REGION Network 7: Send Current Mode
   // Relay current mode to master & slave
   RUNG wire#powerrail
      Move(in := "70_Mode_Data".CRNT_MODE, out1 => "56_SLAVE_CMNDS".CRNT_MODE)
      Move(in := "70_Mode_Data".CRNT_MODE, out1 => "55_STATUS_DATA".CRNT_MODE)
      Move(in := "70_Mode_Data".CRNT_MODE, out1 => "82_To_HMI".CRNT_MODE_IGG)
   END_RUNG
   // the same network as SCL:
   "56_SLAVE_CMNDS".CRNT_MODE := "70_Mode_Data".CRNT_MODE;
   "55_STATUS_DATA".CRNT_MODE := "70_Mode_Data".CRNT_MODE;
   "82_To_HMI".CRNT_MODE_IGG := "70_Mode_Data".CRNT_MODE;
END_REGION

REGION Network 8: Leaving Manual
   // For determination of transition to automatic
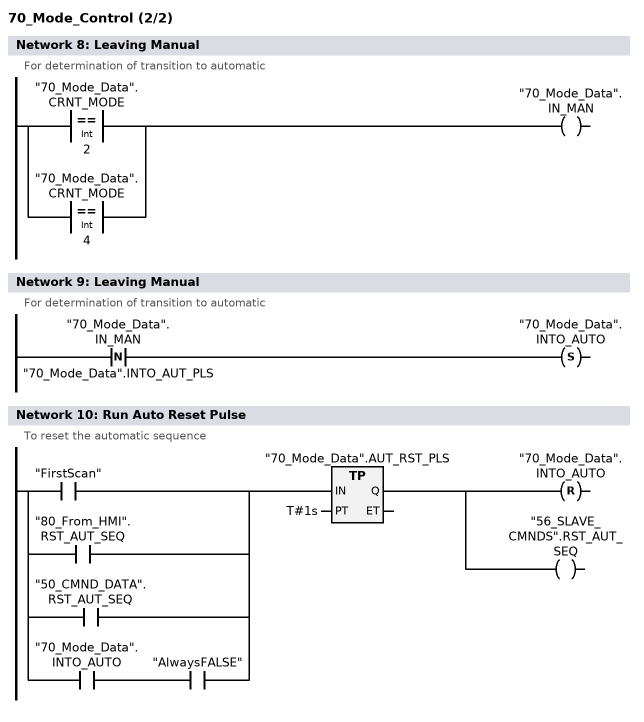
   RUNG wire#powerrail
      { S7_Templates := "SrcType := Int" } EQ_Contact(in1 := "70_Mode_Data".CRNT_MODE, in2 := 2)
      wire#w1
      Coil( "70_Mode_Data".IN_MAN )
   END_RUNG
   RUNG wire#powerrail
      { S7_Templates := "SrcType := Int" } EQ_Contact(in1 := "70_Mode_Data".CRNT_MODE, in2 := 4)
   END_RUNG wire#w1
   // the same network as SCL:
   "70_Mode_Data".IN_MAN := ("70_Mode_Data".CRNT_MODE = 2) OR ("70_Mode_Data".CRNT_MODE = 4);
END_REGION

REGION Network 9: Leaving Manual
   // For determination of transition to automatic
   RUNG wire#powerrail
      N_Contact(operand := "70_Mode_Data".IN_MAN, bit := "70_Mode_Data".INTO_AUT_PLS)
      S_Coil( "70_Mode_Data".INTO_AUTO )
   END_RUNG
   // the same network as SCL:
   #_w1 := NOT "70_Mode_Data".IN_MAN AND "70_Mode_Data".INTO_AUT_PLS;   // falling edge of "70_Mode_Data".IN_MAN
   "70_Mode_Data".INTO_AUT_PLS := "70_Mode_Data".IN_MAN;
   IF #_w1 THEN "70_Mode_Data".INTO_AUTO := TRUE; END_IF;
END_REGION

REGION Network 10: Run Auto Reset Pulse
   // To reset the automatic sequence
   "70_Mode_Data".AUT_RST_PLS.TP(IN := "FirstScan" OR "80_From_HMI".RST_AUT_SEQ OR "50_CMND_DATA".RST_AUT_SEQ OR ("70_Mode_Data".INTO_AUTO AND "AlwaysFALSE"),
                           PT := T#1s);
   IF "70_Mode_Data".AUT_RST_PLS.Q THEN "70_Mode_Data".INTO_AUTO := FALSE; END_IF;
   "56_SLAVE_CMNDS".RST_AUT_SEQ := "70_Mode_Data".AUT_RST_PLS.Q;
END_REGION
END_FUNCTION

// folder: 90 - 99 Manual Functions

FUNCTION_BLOCK "FuelPump"   // FB505, LAD
{ S7_Optimized_Access := 'TRUE' }
VERSION : 0.1
   VAR_INPUT
      Start_Command : Bool;
      Triped : Bool;
      Run : Bool;
      "E-Stop" : Bool;
      Interlock : Bool;
   END_VAR
   VAR_OUTPUT
      Start_Pump : Bool;
   END_VAR
   VAR
      Aux : Struct
         Aux1 : Bool;
         Aux2 : Bool;
      END_STRUCT;
   END_VAR
   VAR_TEMP   // added for the SCL form of the ladder/FBD networks
      _w1 : Bool;
      _w2 : Bool;
      _w3 : Bool;
   END_VAR
BEGIN

REGION Network 1
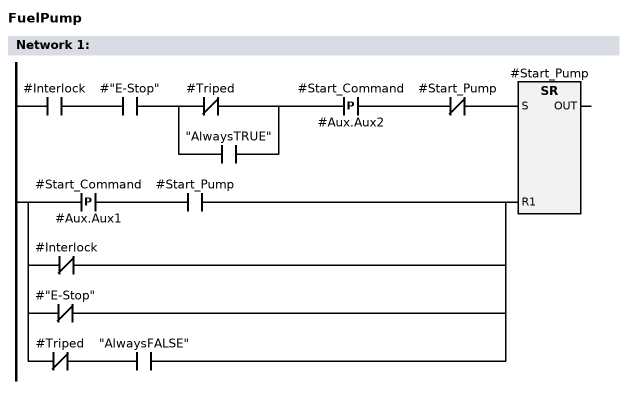
   RUNG wire#powerrail
      Contact( #Interlock )
      Contact( #"E-Stop" )
      wire#w1
      I_Contact( #Triped )
      wire#w2
      P_Contact(operand := #Start_Command, bit := #Aux.Aux2)
      I_Contact( #Start_Pump )
      S_SR(operand := #Start_Pump, r1 := wire#w3)
   END_RUNG
   RUNG wire#w1
      Contact( "AlwaysTRUE" )
   END_RUNG wire#w2
   RUNG wire#powerrail
      P_Contact(operand := #Start_Command, bit := #Aux.Aux1)
      Contact( #Start_Pump )
   END_RUNG wire#w3
   RUNG wire#powerrail
      I_Contact( #Interlock )
   END_RUNG wire#w3
   RUNG wire#powerrail
      I_Contact( #"E-Stop" )
   END_RUNG wire#w3
   RUNG wire#powerrail
      I_Contact( #Triped )
      Contact( "AlwaysFALSE" )
   END_RUNG wire#w3
   // the same network as SCL:
   #_w1 := #Interlock AND #"E-Stop" AND (NOT #Triped OR "AlwaysTRUE") AND #Start_Command AND NOT #Aux.Aux2;   // rising edge of #Start_Command
   #Aux.Aux2 := #Start_Command;
   #_w2 := #Start_Command AND NOT #Aux.Aux1;   // rising edge of #Start_Command
   #Aux.Aux1 := #Start_Command;
   #_w3 := (#_w2 AND #Start_Pump) OR NOT #Interlock OR NOT #"E-Stop" OR (NOT #Triped AND "AlwaysFALSE");
   IF #_w1 AND NOT #Start_Pump THEN
       #Start_Pump := TRUE;   // SR flip-flop
   END_IF;
   IF #_w3 THEN #Start_Pump := FALSE; END_IF;
END_REGION
END_FUNCTION_BLOCK

FUNCTION "90_Manual_Control" : Void   // FC90, LAD
TITLE = Manual Control
{ S7_Optimized_Access := 'TRUE' }
AUTHOR : JHT
VERSION : 0.1
// Code for manual operation of equipment
   VAR_TEMP
      Aux : Struct
         Aux1 : Bool;
      END_STRUCT;
   END_VAR
   VAR_TEMP   // added for the SCL form of the ladder/FBD networks
      _w1 : Bool;
      _w2 : Bool;
      _w3 : Bool;
      _w4 : Bool;
      _w5 : Bool;
      _w6 : Bool;
   END_VAR
BEGIN

REGION Network 1: Zero Auto Step Numbers
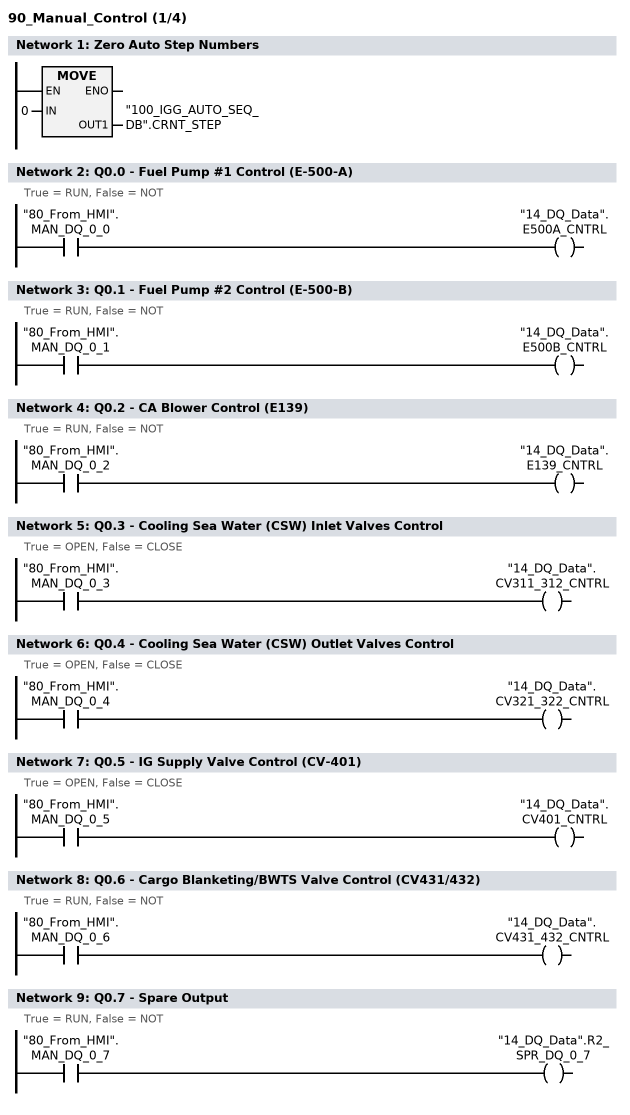
   RUNG wire#powerrail
      Move(in := 0, out1 => "100_IGG_AUTO_SEQ_DB".CRNT_STEP)
   END_RUNG
   // the same network as SCL:
   "100_IGG_AUTO_SEQ_DB".CRNT_STEP := 0;
END_REGION

REGION Network 2: Q0.0 - Fuel Pump #1 Control (E-500-A)
   // True = RUN, False = NOT
   RUNG wire#powerrail
      Contact( "80_From_HMI".MAN_DQ_0_0 )
      Coil( "14_DQ_Data".E500A_CNTRL )
   END_RUNG
   // the same network as SCL:
   "14_DQ_Data".E500A_CNTRL := "80_From_HMI".MAN_DQ_0_0;
END_REGION

REGION Network 3: Q0.1 - Fuel Pump #2 Control (E-500-B)
   // True = RUN, False = NOT
   RUNG wire#powerrail
      Contact( "80_From_HMI".MAN_DQ_0_1 )
      Coil( "14_DQ_Data".E500B_CNTRL )
   END_RUNG
   // the same network as SCL:
   "14_DQ_Data".E500B_CNTRL := "80_From_HMI".MAN_DQ_0_1;
END_REGION

REGION Network 4: Q0.2 - CA Blower Control (E139)
   // True = RUN, False = NOT
   RUNG wire#powerrail
      Contact( "80_From_HMI".MAN_DQ_0_2 )
      Coil( "14_DQ_Data".E139_CNTRL )
   END_RUNG
   // the same network as SCL:
   "14_DQ_Data".E139_CNTRL := "80_From_HMI".MAN_DQ_0_2;
END_REGION

REGION Network 5: Q0.3 - Cooling Sea Water (CSW) Inlet Valves Control
   // True = OPEN, False = CLOSE
   RUNG wire#powerrail
      Contact( "80_From_HMI".MAN_DQ_0_3 )
      Coil( "14_DQ_Data".CV311_312_CNTRL )
   END_RUNG
   // the same network as SCL:
   "14_DQ_Data".CV311_312_CNTRL := "80_From_HMI".MAN_DQ_0_3;
END_REGION

REGION Network 6: Q0.4 - Cooling Sea Water (CSW) Outlet Valves Control
   // True = OPEN, False = CLOSE
   RUNG wire#powerrail
      Contact( "80_From_HMI".MAN_DQ_0_4 )
      Coil( "14_DQ_Data".CV321_322_CNTRL )
   END_RUNG
   // the same network as SCL:
   "14_DQ_Data".CV321_322_CNTRL := "80_From_HMI".MAN_DQ_0_4;
END_REGION

REGION Network 7: Q0.5 - IG Supply Valve Control (CV-401)
   // True = OPEN, False = CLOSE
   RUNG wire#powerrail
      Contact( "80_From_HMI".MAN_DQ_0_5 )
      Coil( "14_DQ_Data".CV401_CNTRL )
   END_RUNG
   // the same network as SCL:
   "14_DQ_Data".CV401_CNTRL := "80_From_HMI".MAN_DQ_0_5;
END_REGION

REGION Network 8: Q0.6 - Cargo Blanketing/BWTS Valve Control (CV431/432)
   // True = RUN, False = NOT
   RUNG wire#powerrail
      Contact( "80_From_HMI".MAN_DQ_0_6 )
      Coil( "14_DQ_Data".CV431_432_CNTRL )
   END_RUNG
   // the same network as SCL:
   "14_DQ_Data".CV431_432_CNTRL := "80_From_HMI".MAN_DQ_0_6;
END_REGION

REGION Network 9: Q0.7 - Spare Output
   // True = RUN, False = NOT
   RUNG wire#powerrail
      Contact( "80_From_HMI".MAN_DQ_0_7 )
      Coil( "14_DQ_Data".R2_SPR_DQ_0_7 )
   END_RUNG
   // the same network as SCL:
   "14_DQ_Data".R2_SPR_DQ_0_7 := "80_From_HMI".MAN_DQ_0_7;
END_REGION

REGION Network 10: Q1.0 - Spare Output
   // True = RUN, False = NOT
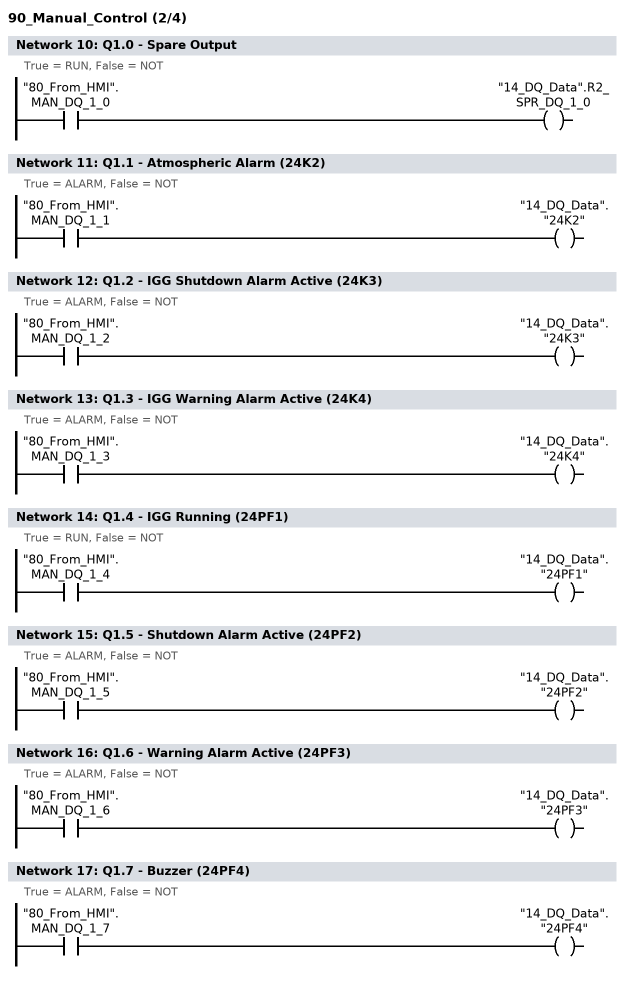
   RUNG wire#powerrail
      Contact( "80_From_HMI".MAN_DQ_1_0 )
      Coil( "14_DQ_Data".R2_SPR_DQ_1_0 )
   END_RUNG
   // the same network as SCL:
   "14_DQ_Data".R2_SPR_DQ_1_0 := "80_From_HMI".MAN_DQ_1_0;
END_REGION

REGION Network 11: Q1.1 - Atmospheric Alarm (24K2)
   // True = ALARM, False = NOT
   RUNG wire#powerrail
      Contact( "80_From_HMI".MAN_DQ_1_1 )
      Coil( "14_DQ_Data"."24K2" )
   END_RUNG
   // the same network as SCL:
   "14_DQ_Data"."24K2" := "80_From_HMI".MAN_DQ_1_1;
END_REGION

REGION Network 12: Q1.2 - IGG Shutdown Alarm Active (24K3)
   // True = ALARM, False = NOT
   RUNG wire#powerrail
      Contact( "80_From_HMI".MAN_DQ_1_2 )
      Coil( "14_DQ_Data"."24K3" )
   END_RUNG
   // the same network as SCL:
   "14_DQ_Data"."24K3" := "80_From_HMI".MAN_DQ_1_2;
END_REGION

REGION Network 13: Q1.3 - IGG Warning Alarm Active (24K4)
   // True = ALARM, False = NOT
   RUNG wire#powerrail
      Contact( "80_From_HMI".MAN_DQ_1_3 )
      Coil( "14_DQ_Data"."24K4" )
   END_RUNG
   // the same network as SCL:
   "14_DQ_Data"."24K4" := "80_From_HMI".MAN_DQ_1_3;
END_REGION

REGION Network 14: Q1.4 - IGG Running (24PF1)
   // True = RUN, False = NOT
   RUNG wire#powerrail
      Contact( "80_From_HMI".MAN_DQ_1_4 )
      Coil( "14_DQ_Data"."24PF1" )
   END_RUNG
   // the same network as SCL:
   "14_DQ_Data"."24PF1" := "80_From_HMI".MAN_DQ_1_4;
END_REGION

REGION Network 15: Q1.5 - Shutdown Alarm Active (24PF2)
   // True = ALARM, False = NOT
   RUNG wire#powerrail
      Contact( "80_From_HMI".MAN_DQ_1_5 )
      Coil( "14_DQ_Data"."24PF2" )
   END_RUNG
   // the same network as SCL:
   "14_DQ_Data"."24PF2" := "80_From_HMI".MAN_DQ_1_5;
END_REGION

REGION Network 16: Q1.6 - Warning Alarm Active (24PF3)
   // True = ALARM, False = NOT
   RUNG wire#powerrail
      Contact( "80_From_HMI".MAN_DQ_1_6 )
      Coil( "14_DQ_Data"."24PF3" )
   END_RUNG
   // the same network as SCL:
   "14_DQ_Data"."24PF3" := "80_From_HMI".MAN_DQ_1_6;
END_REGION

REGION Network 17: Q1.7 - Buzzer (24PF4)
   // True = ALARM, False = NOT
   RUNG wire#powerrail
      Contact( "80_From_HMI".MAN_DQ_1_7 )
      Coil( "14_DQ_Data"."24PF4" )
   END_RUNG
   // the same network as SCL:
   "14_DQ_Data"."24PF4" := "80_From_HMI".MAN_DQ_1_7;
END_REGION

REGION Network 18: QW98 - Vent Valve Position Control (CV-403)
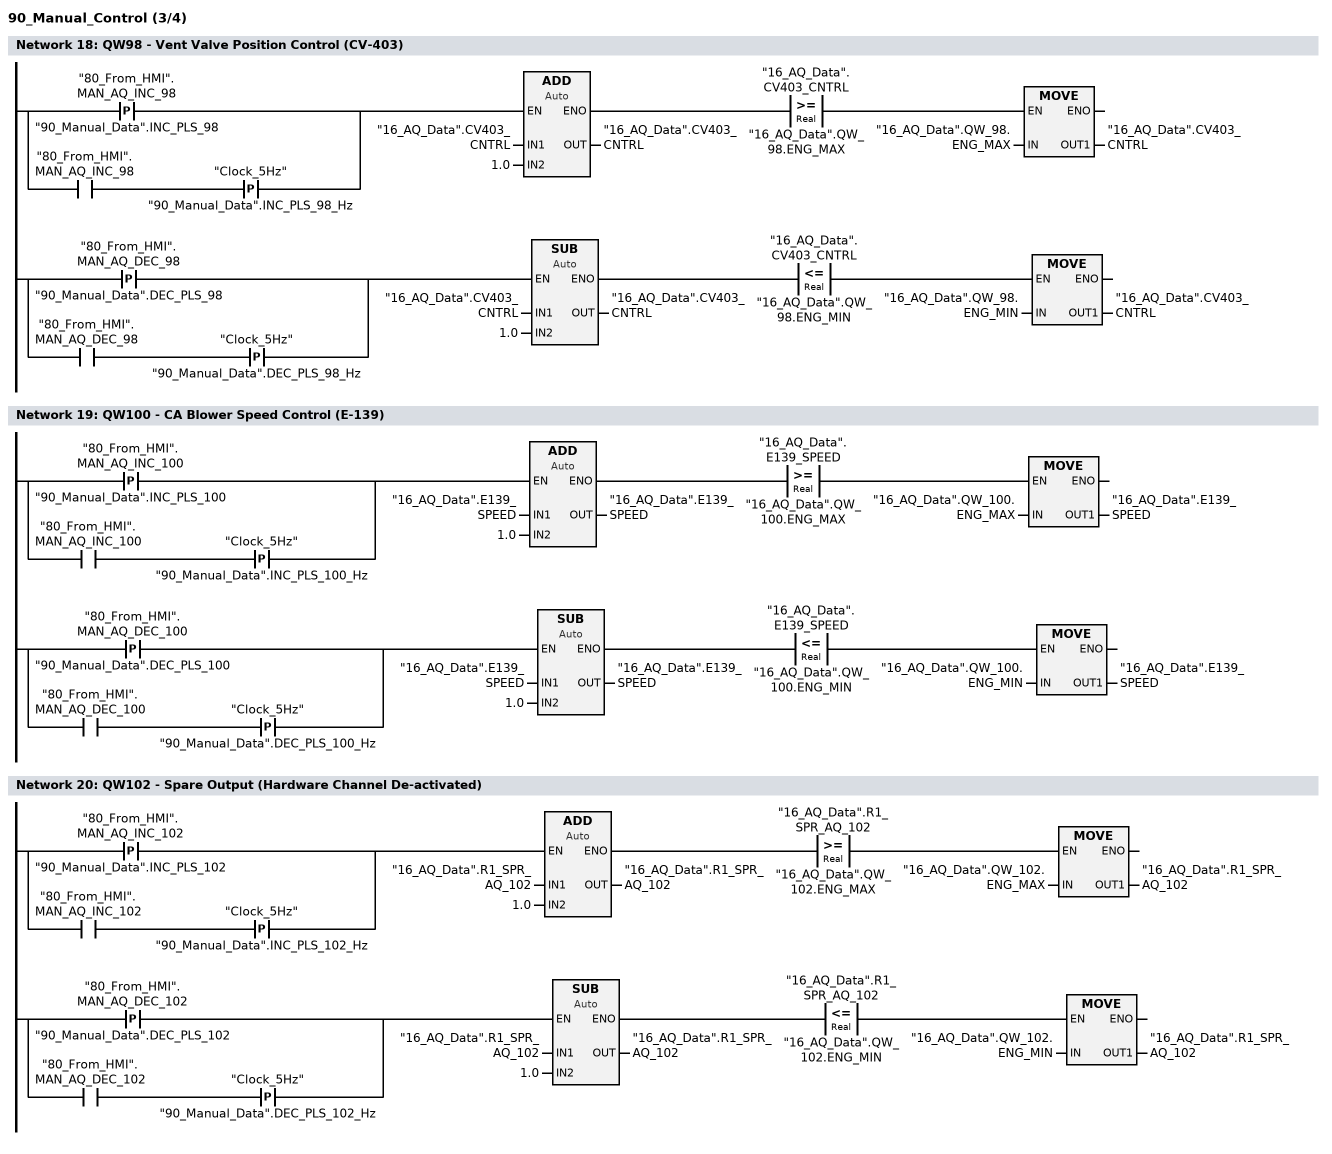
   RUNG wire#powerrail
      P_Contact(operand := "80_From_HMI".MAN_AQ_INC_98, bit := "90_Manual_Data".INC_PLS_98)
      wire#w1
      Add(in1 := "16_AQ_Data".CV403_CNTRL, in2 := 1.0, out => "16_AQ_Data".CV403_CNTRL)
      { S7_Templates := "SrcType := Real" } GE_Contact(in1 := "16_AQ_Data".CV403_CNTRL, in2 := "16_AQ_Data".QW_98.ENG_MAX)
      { S7_GenerateENO := "TRUE" } Move(in := "16_AQ_Data".QW_98.ENG_MAX, out1 => "16_AQ_Data".CV403_CNTRL)
   END_RUNG
   RUNG wire#powerrail
      Contact( "80_From_HMI".MAN_AQ_INC_98 )
      P_Contact(operand := "Clock_5Hz", bit := "90_Manual_Data".INC_PLS_98_Hz)
   END_RUNG wire#w1
   RUNG wire#powerrail
      P_Contact(operand := "80_From_HMI".MAN_AQ_DEC_98, bit := "90_Manual_Data".DEC_PLS_98)
      wire#w2
      Sub(in1 := "16_AQ_Data".CV403_CNTRL, in2 := 1.0, out => "16_AQ_Data".CV403_CNTRL)
      { S7_Templates := "SrcType := Real" } LE_Contact(in1 := "16_AQ_Data".CV403_CNTRL, in2 := "16_AQ_Data".QW_98.ENG_MIN)
      { S7_GenerateENO := "TRUE" } Move(in := "16_AQ_Data".QW_98.ENG_MIN, out1 => "16_AQ_Data".CV403_CNTRL)
   END_RUNG
   RUNG wire#powerrail
      Contact( "80_From_HMI".MAN_AQ_DEC_98 )
      P_Contact(operand := "Clock_5Hz", bit := "90_Manual_Data".DEC_PLS_98_Hz)
   END_RUNG wire#w2
   // the same network as SCL:
   #_w1 := "80_From_HMI".MAN_AQ_INC_98 AND NOT "90_Manual_Data".INC_PLS_98;   // rising edge of "80_From_HMI".MAN_AQ_INC_98
   "90_Manual_Data".INC_PLS_98 := "80_From_HMI".MAN_AQ_INC_98;
   #_w2 := "80_From_HMI".MAN_AQ_INC_98 AND "Clock_5Hz" AND NOT "90_Manual_Data".INC_PLS_98_Hz;   // rising edge of "Clock_5Hz"
   "90_Manual_Data".INC_PLS_98_Hz := "Clock_5Hz";
   #_w3 := #_w1 OR #_w2;
   IF #_w3 THEN "16_AQ_Data".CV403_CNTRL := "16_AQ_Data".CV403_CNTRL + 1.0; END_IF;
   IF #_w3 AND ("16_AQ_Data".CV403_CNTRL >= "16_AQ_Data".QW_98.ENG_MAX) THEN
       "16_AQ_Data".CV403_CNTRL := "16_AQ_Data".QW_98.ENG_MAX;
   END_IF;
   #_w4 := "80_From_HMI".MAN_AQ_DEC_98 AND NOT "90_Manual_Data".DEC_PLS_98;   // rising edge of "80_From_HMI".MAN_AQ_DEC_98
   "90_Manual_Data".DEC_PLS_98 := "80_From_HMI".MAN_AQ_DEC_98;
   #_w5 := "80_From_HMI".MAN_AQ_DEC_98 AND "Clock_5Hz" AND NOT "90_Manual_Data".DEC_PLS_98_Hz;   // rising edge of "Clock_5Hz"
   "90_Manual_Data".DEC_PLS_98_Hz := "Clock_5Hz";
   #_w6 := #_w4 OR #_w5;
   IF #_w6 THEN "16_AQ_Data".CV403_CNTRL := "16_AQ_Data".CV403_CNTRL - 1.0; END_IF;
   IF #_w6 AND ("16_AQ_Data".CV403_CNTRL <= "16_AQ_Data".QW_98.ENG_MIN) THEN
       "16_AQ_Data".CV403_CNTRL := "16_AQ_Data".QW_98.ENG_MIN;
   END_IF;
END_REGION

REGION Network 19: QW100 - CA Blower Speed Control (E-139)
   RUNG wire#powerrail
      P_Contact(operand := "80_From_HMI".MAN_AQ_INC_100, bit := "90_Manual_Data".INC_PLS_100)
      wire#w1
      Add(in1 := "16_AQ_Data".E139_SPEED, in2 := 1.0, out => "16_AQ_Data".E139_SPEED)
      { S7_Templates := "SrcType := Real" } GE_Contact(in1 := "16_AQ_Data".E139_SPEED, in2 := "16_AQ_Data".QW_100.ENG_MAX)
      { S7_GenerateENO := "TRUE" } Move(in := "16_AQ_Data".QW_100.ENG_MAX, out1 => "16_AQ_Data".E139_SPEED)
   END_RUNG
   RUNG wire#powerrail
      Contact( "80_From_HMI".MAN_AQ_INC_100 )
      P_Contact(operand := "Clock_5Hz", bit := "90_Manual_Data".INC_PLS_100_Hz)
   END_RUNG wire#w1
   RUNG wire#powerrail
      P_Contact(operand := "80_From_HMI".MAN_AQ_DEC_100, bit := "90_Manual_Data".DEC_PLS_100)
      wire#w2
      Sub(in1 := "16_AQ_Data".E139_SPEED, in2 := 1.0, out => "16_AQ_Data".E139_SPEED)
      { S7_Templates := "SrcType := Real" } LE_Contact(in1 := "16_AQ_Data".E139_SPEED, in2 := "16_AQ_Data".QW_100.ENG_MIN)
      { S7_GenerateENO := "TRUE" } Move(in := "16_AQ_Data".QW_100.ENG_MIN, out1 => "16_AQ_Data".E139_SPEED)
   END_RUNG
   RUNG wire#powerrail
      Contact( "80_From_HMI".MAN_AQ_DEC_100 )
      P_Contact(operand := "Clock_5Hz", bit := "90_Manual_Data".DEC_PLS_100_Hz)
   END_RUNG wire#w2
   // the same network as SCL:
   #_w1 := "80_From_HMI".MAN_AQ_INC_100 AND NOT "90_Manual_Data".INC_PLS_100;   // rising edge of "80_From_HMI".MAN_AQ_INC_100
   "90_Manual_Data".INC_PLS_100 := "80_From_HMI".MAN_AQ_INC_100;
   #_w2 := "80_From_HMI".MAN_AQ_INC_100 AND "Clock_5Hz" AND NOT "90_Manual_Data".INC_PLS_100_Hz;   // rising edge of "Clock_5Hz"
   "90_Manual_Data".INC_PLS_100_Hz := "Clock_5Hz";
   #_w3 := #_w1 OR #_w2;
   IF #_w3 THEN "16_AQ_Data".E139_SPEED := "16_AQ_Data".E139_SPEED + 1.0; END_IF;
   IF #_w3 AND ("16_AQ_Data".E139_SPEED >= "16_AQ_Data".QW_100.ENG_MAX) THEN
       "16_AQ_Data".E139_SPEED := "16_AQ_Data".QW_100.ENG_MAX;
   END_IF;
   #_w4 := "80_From_HMI".MAN_AQ_DEC_100 AND NOT "90_Manual_Data".DEC_PLS_100;   // rising edge of "80_From_HMI".MAN_AQ_DEC_100
   "90_Manual_Data".DEC_PLS_100 := "80_From_HMI".MAN_AQ_DEC_100;
   #_w5 := "80_From_HMI".MAN_AQ_DEC_100 AND "Clock_5Hz" AND NOT "90_Manual_Data".DEC_PLS_100_Hz;   // rising edge of "Clock_5Hz"
   "90_Manual_Data".DEC_PLS_100_Hz := "Clock_5Hz";
   #_w6 := #_w4 OR #_w5;
   IF #_w6 THEN "16_AQ_Data".E139_SPEED := "16_AQ_Data".E139_SPEED - 1.0; END_IF;
   IF #_w6 AND ("16_AQ_Data".E139_SPEED <= "16_AQ_Data".QW_100.ENG_MIN) THEN
       "16_AQ_Data".E139_SPEED := "16_AQ_Data".QW_100.ENG_MIN;
   END_IF;
END_REGION

REGION Network 20: QW102 - Spare Output (Hardware Channel De-activated)
   RUNG wire#powerrail
      P_Contact(operand := "80_From_HMI".MAN_AQ_INC_102, bit := "90_Manual_Data".INC_PLS_102)
      wire#w1
      Add(in1 := "16_AQ_Data".R1_SPR_AQ_102, in2 := 1.0, out => "16_AQ_Data".R1_SPR_AQ_102)
      { S7_Templates := "SrcType := Real" } GE_Contact(in1 := "16_AQ_Data".R1_SPR_AQ_102, in2 := "16_AQ_Data".QW_102.ENG_MAX)
      { S7_GenerateENO := "TRUE" } Move(in := "16_AQ_Data".QW_102.ENG_MAX, out1 => "16_AQ_Data".R1_SPR_AQ_102)
   END_RUNG
   RUNG wire#powerrail
      Contact( "80_From_HMI".MAN_AQ_INC_102 )
      P_Contact(operand := "Clock_5Hz", bit := "90_Manual_Data".INC_PLS_102_Hz)
   END_RUNG wire#w1
   RUNG wire#powerrail
      P_Contact(operand := "80_From_HMI".MAN_AQ_DEC_102, bit := "90_Manual_Data".DEC_PLS_102)
      wire#w2
      Sub(in1 := "16_AQ_Data".R1_SPR_AQ_102, in2 := 1.0, out => "16_AQ_Data".R1_SPR_AQ_102)
      { S7_Templates := "SrcType := Real" } LE_Contact(in1 := "16_AQ_Data".R1_SPR_AQ_102, in2 := "16_AQ_Data".QW_102.ENG_MIN)
      { S7_GenerateENO := "TRUE" } Move(in := "16_AQ_Data".QW_102.ENG_MIN, out1 => "16_AQ_Data".R1_SPR_AQ_102)
   END_RUNG
   RUNG wire#powerrail
      Contact( "80_From_HMI".MAN_AQ_DEC_102 )
      P_Contact(operand := "Clock_5Hz", bit := "90_Manual_Data".DEC_PLS_102_Hz)
   END_RUNG wire#w2
   // the same network as SCL:
   #_w1 := "80_From_HMI".MAN_AQ_INC_102 AND NOT "90_Manual_Data".INC_PLS_102;   // rising edge of "80_From_HMI".MAN_AQ_INC_102
   "90_Manual_Data".INC_PLS_102 := "80_From_HMI".MAN_AQ_INC_102;
   #_w2 := "80_From_HMI".MAN_AQ_INC_102 AND "Clock_5Hz" AND NOT "90_Manual_Data".INC_PLS_102_Hz;   // rising edge of "Clock_5Hz"
   "90_Manual_Data".INC_PLS_102_Hz := "Clock_5Hz";
   #_w3 := #_w1 OR #_w2;
   IF #_w3 THEN "16_AQ_Data".R1_SPR_AQ_102 := "16_AQ_Data".R1_SPR_AQ_102 + 1.0; END_IF;
   IF #_w3 AND ("16_AQ_Data".R1_SPR_AQ_102 >= "16_AQ_Data".QW_102.ENG_MAX) THEN
       "16_AQ_Data".R1_SPR_AQ_102 := "16_AQ_Data".QW_102.ENG_MAX;
   END_IF;
   #_w4 := "80_From_HMI".MAN_AQ_DEC_102 AND NOT "90_Manual_Data".DEC_PLS_102;   // rising edge of "80_From_HMI".MAN_AQ_DEC_102
   "90_Manual_Data".DEC_PLS_102 := "80_From_HMI".MAN_AQ_DEC_102;
   #_w5 := "80_From_HMI".MAN_AQ_DEC_102 AND "Clock_5Hz" AND NOT "90_Manual_Data".DEC_PLS_102_Hz;   // rising edge of "Clock_5Hz"
   "90_Manual_Data".DEC_PLS_102_Hz := "Clock_5Hz";
   #_w6 := #_w4 OR #_w5;
   IF #_w6 THEN "16_AQ_Data".R1_SPR_AQ_102 := "16_AQ_Data".R1_SPR_AQ_102 - 1.0; END_IF;
   IF #_w6 AND ("16_AQ_Data".R1_SPR_AQ_102 <= "16_AQ_Data".QW_102.ENG_MIN) THEN
       "16_AQ_Data".R1_SPR_AQ_102 := "16_AQ_Data".QW_102.ENG_MIN;
   END_IF;
END_REGION

REGION Network 21: QW104 - Spare Output (Hardware Channel De-activated)
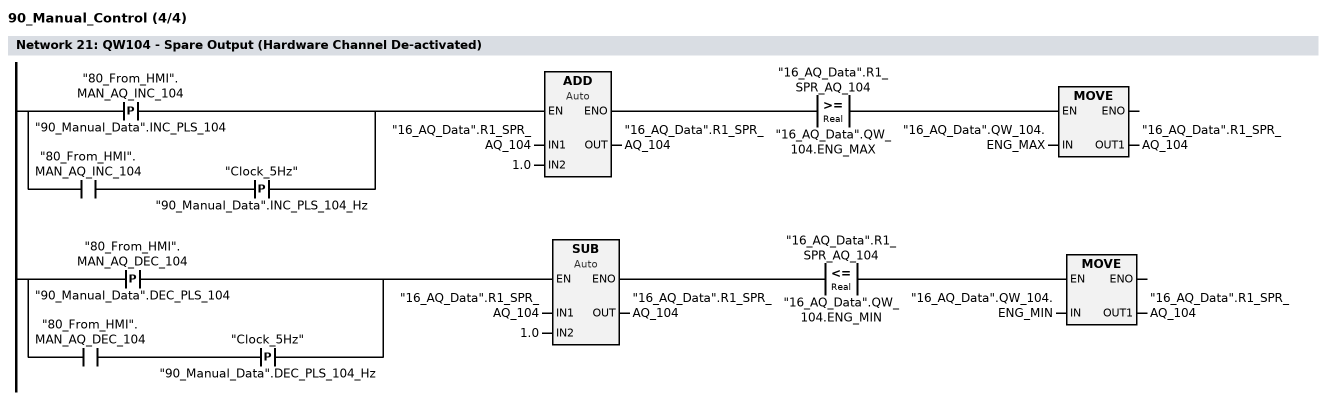
   RUNG wire#powerrail
      P_Contact(operand := "80_From_HMI".MAN_AQ_INC_104, bit := "90_Manual_Data".INC_PLS_104)
      wire#w1
      Add(in1 := "16_AQ_Data".R1_SPR_AQ_104, in2 := 1.0, out => "16_AQ_Data".R1_SPR_AQ_104)
      { S7_Templates := "SrcType := Real" } GE_Contact(in1 := "16_AQ_Data".R1_SPR_AQ_104, in2 := "16_AQ_Data".QW_104.ENG_MAX)
      { S7_GenerateENO := "TRUE" } Move(in := "16_AQ_Data".QW_104.ENG_MAX, out1 => "16_AQ_Data".R1_SPR_AQ_104)
   END_RUNG
   RUNG wire#powerrail
      Contact( "80_From_HMI".MAN_AQ_INC_104 )
      P_Contact(operand := "Clock_5Hz", bit := "90_Manual_Data".INC_PLS_104_Hz)
   END_RUNG wire#w1
   RUNG wire#powerrail
      P_Contact(operand := "80_From_HMI".MAN_AQ_DEC_104, bit := "90_Manual_Data".DEC_PLS_104)
      wire#w2
      Sub(in1 := "16_AQ_Data".R1_SPR_AQ_104, in2 := 1.0, out => "16_AQ_Data".R1_SPR_AQ_104)
      { S7_Templates := "SrcType := Real" } LE_Contact(in1 := "16_AQ_Data".R1_SPR_AQ_104, in2 := "16_AQ_Data".QW_104.ENG_MIN)
      { S7_GenerateENO := "TRUE" } Move(in := "16_AQ_Data".QW_104.ENG_MIN, out1 => "16_AQ_Data".R1_SPR_AQ_104)
   END_RUNG
   RUNG wire#powerrail
      Contact( "80_From_HMI".MAN_AQ_DEC_104 )
      P_Contact(operand := "Clock_5Hz", bit := "90_Manual_Data".DEC_PLS_104_Hz)
   END_RUNG wire#w2
   // the same network as SCL:
   #_w1 := "80_From_HMI".MAN_AQ_INC_104 AND NOT "90_Manual_Data".INC_PLS_104;   // rising edge of "80_From_HMI".MAN_AQ_INC_104
   "90_Manual_Data".INC_PLS_104 := "80_From_HMI".MAN_AQ_INC_104;
   #_w2 := "80_From_HMI".MAN_AQ_INC_104 AND "Clock_5Hz" AND NOT "90_Manual_Data".INC_PLS_104_Hz;   // rising edge of "Clock_5Hz"
   "90_Manual_Data".INC_PLS_104_Hz := "Clock_5Hz";
   #_w3 := #_w1 OR #_w2;
   IF #_w3 THEN "16_AQ_Data".R1_SPR_AQ_104 := "16_AQ_Data".R1_SPR_AQ_104 + 1.0; END_IF;
   IF #_w3 AND ("16_AQ_Data".R1_SPR_AQ_104 >= "16_AQ_Data".QW_104.ENG_MAX) THEN
       "16_AQ_Data".R1_SPR_AQ_104 := "16_AQ_Data".QW_104.ENG_MAX;
   END_IF;
   #_w4 := "80_From_HMI".MAN_AQ_DEC_104 AND NOT "90_Manual_Data".DEC_PLS_104;   // rising edge of "80_From_HMI".MAN_AQ_DEC_104
   "90_Manual_Data".DEC_PLS_104 := "80_From_HMI".MAN_AQ_DEC_104;
   #_w5 := "80_From_HMI".MAN_AQ_DEC_104 AND "Clock_5Hz" AND NOT "90_Manual_Data".DEC_PLS_104_Hz;   // rising edge of "Clock_5Hz"
   "90_Manual_Data".DEC_PLS_104_Hz := "Clock_5Hz";
   #_w6 := #_w4 OR #_w5;
   IF #_w6 THEN "16_AQ_Data".R1_SPR_AQ_104 := "16_AQ_Data".R1_SPR_AQ_104 - 1.0; END_IF;
   IF #_w6 AND ("16_AQ_Data".R1_SPR_AQ_104 <= "16_AQ_Data".QW_104.ENG_MIN) THEN
       "16_AQ_Data".R1_SPR_AQ_104 := "16_AQ_Data".QW_104.ENG_MIN;
   END_IF;
END_REGION
END_FUNCTION

// ===== PLC "Rack 2 - BC PLC - 15KF3"  CPU 1510SP-1 PN =====

VAR_GLOBAL   // PLC tag table "Default tag table"
   "System_Byte" AT %MB1 : Byte;
   "FirstScan" AT %M1.0 : Bool;
   "DiagStatusUpdate" AT %M1.1 : Bool;
   "AlwaysTRUE" AT %M1.2 : Bool;
   "AlwaysFALSE" AT %M1.3 : Bool;
   "Clock_Byte" AT %MB0 : Byte;
   "Clock_10Hz" AT %M0.0 : Bool;
   "Clock_5Hz" AT %M0.1 : Bool;
   "Clock_2.5Hz" AT %M0.2 : Bool;
   "Clock_2Hz" AT %M0.3 : Bool;
   "Clock_1.25Hz" AT %M0.4 : Bool;
   "Clock_1Hz" AT %M0.5 : Bool;
   "Clock_0.625Hz" AT %M0.6 : Bool;
   "Clock_0.5Hz" AT %M0.7 : Bool;
   "CA Pressure Switch (PS101)" AT %I0.0 : Bool;   // PS101-19B1
   "IA Compressor Shutdown" AT %I0.1 : Bool;   // E131-MCCP/IA-Comp
   "R1_SPR_DI_0_2" AT %I0.2 : Bool;   // Spare Input
   "R1_SPR_DI_0_3" AT %I0.3 : Bool;   // Spare input
   "Igniter Power Healthy" AT %I0.4 : Bool;   // X001-6Q6
   "FDU Power Healthy" AT %I0.5 : Bool;   // FD001-6Q5
   "FDU Healthy" AT %I0.6 : Bool;   // FD001-9K1
   "Burner Flame Detected" AT %I0.7 : Bool;   // FD001-9BR1
   "Pilot Ignition Air Flow Switch" AT %I1.0 : Bool;   // FS123-20B1
   "Main Atom Air Flow Switch" AT %I1.1 : Bool;   // FS115-20B2
   "Nozzle Cooling Water Flow Switch" AT %I1.2 : Bool;   // FS320-20B3
   "Jacket Cooling Water Flow Switch" AT %I1.3 : Bool;   // FS317-20B4
   "CSW Pump Tripped" AT %I1.4 : Bool;   // P301-MCCP/7Q5
   "CSW Pump Enabled" AT %I1.5 : Bool;   // P301-MCCP/12Q1
   "External Shutdown" AT %I1.7 : Bool;   // ESD
   "O2 Analyser System Fail" AT %I2.0 : Bool;   // E600-11B1
   "O2 Analyser Hi Hi" AT %I2.1 : Bool;   // E600-11B1
   "O2 Analyser Lo Lo" AT %I2.2 : Bool;   // E600-11B1
   "O2 System Power Healthy" AT %I2.3 : Bool;   // E600-6Q7
   "Soot System Power Healthy" AT %I2.4 : Bool;   // E700-6Q8
   "Soot System Opacity" AT %I2.5 : Bool;   // E700-12B1
   "IG Temp Hi Hi Switch" AT %I2.6 : Bool;   // TS403-21K1
   "IG Shell Temp Hi Switch" AT %I2.7 : Bool;   // TS006--21K2
   "IGG E-Stop Healthy" AT %I3.0 : Bool;   // S2-8K1
   "IA Comp Warning" AT %I3.1 : Bool;   // E131-MCCP/IA-Comp
   "R2_SPR_DI_3_2" AT %I3.2 : Bool;   // Spare Input
   "IA Comp Healthy" AT %I3.3 : Bool;   // E131-MCCP/IA-Comp
   "Shell CW Level Hi Hi Switch" AT %I3.4 : Bool;   // LS001-22B1
   "Fresh Water Pump Tripped" AT %I3.5 : Bool;   // P305
   "Fresh Water Pump Enabled" AT %I3.6 : Bool;   // P305
   "R2_SPR_DI_3_7" AT %I3.7 : Bool;   // Spare input
   "IGG Main Atom Air Pressure" AT %IW100 : Int;   // PIT113-33B2
   "IGG Inlet Fuel Pressure" AT %IW104 : Int;   // PIT204-34B1
   "IGG Inlet Fuel Temp" AT %IW106 : Int;   // TIT202-34B2
   "O2 Analyser Content" AT %IW108 : Int;   // E600-11B1
   "IG Soot Content" AT %IW110 : Int;   // E700-12B1
   "IGG Main Fuel Pressure" AT %IW96 : Int;   // PIT205-33B1
   "Flame Signal" AT %IW98 : Int;   // FD001-9BR1
   "Test Pressure Valve Control" AT %Q0.0 : Bool;   // CV127-25QM1
   "Pilot B Ignition Air Valve Control" AT %Q0.1 : Bool;   // CV124-25QM2
   "Pilot B Fuel Valve 1 Control" AT %Q0.2 : Bool;   // CV215-25QM3
   "Pilot B Fuel Valve 2 Control" AT %Q0.3 : Bool;   // CV216-25QM4
   "Main B Atom Air Valve Control" AT %Q0.4 : Bool;   // CV114-25QM5
   "Main B Fuel Valve 1 Control" AT %Q0.5 : Bool;   // CV206-25QM6
   "Main B Fuel Valve 2 Control" AT %Q0.6 : Bool;   // CV207-25QM7
   "IA Comp Control" AT %Q0.7 : Bool;   // E131-MCCP/IA-Comp
   "CSW Pump Control" AT %Q1.0 : Bool;   // P301-24K1
   "Igniter Control" AT %Q1.1 : Bool;   // X001-27K1
   "R2_SPR_DQ_1_2" AT %Q1.2 : Bool;   // Spare output
   "R2_SPR_DQ_1_3" AT %Q1.3 : Bool;   // Spare output
   "R2_SPR_DQ_1_4" AT %Q1.4 : Bool;   // Spare output
   "R2_SPR_DQ_1_5" AT %Q1.5 : Bool;   // Spare output
   "R2_SPR_DQ_1_6" AT %Q1.6 : Bool;   // Spare output
   "Fresh Water Pump Control" AT %Q1.7 : Bool;   // P305
   "Main Fuel Reg Valve Control" AT %QW100 : Int;   // CV203-38QN1
   "Main Atom Air Reg Valve Control" AT %QW102 : Int;   // CV111-38QN2
   "R2_SPR_AQ_96" AT %QW96 : Int;   // Spare output
   "R2_SPR_DI_1_6" AT %I1.6 : Bool;   // Spare input
   "Inlet IA Pressure PIT112" AT %IW102 : Int;   // PIT112-31B3
   "R2_SPR_AQ_98" AT %QW98 : Int;   // Spare output
   "Test 1" AT %QD104 : Real;
   "LevelBetter" AT %Q108.0 : Bool;
   "IA Comp Healthy/Running" AT %I3.3 : Bool;   // E131-MCCP/IA-Comp
   "Tag_1" AT %M15.0 : Bool;
END_VAR

TYPE "AI_Data"
VERSION : 0.1
   STRUCT
      RAW_MIN : Int;   // Raw minimum value from AI card
      RAW_MAX : Int := 27648;   // Raw maximum value from AI card
      NORM : Real;   // Normalised real value
      ENG_MIN : Real;   // Engineering units minimum value
      ENG_MAX : Real := 100.0;   // Engineering units maximum value
   END_STRUCT;
END_TYPE

TYPE "AQ_Data"
VERSION : 0.1
   STRUCT
      ENG_MIN : Real;   // Engineering units minimum value
      ENG_MAX : Real := 100.0;   // Engineering units maximum value
      NORM : Real;   // Normalised real value
      RAW_MIN : Int;   // Raw minimum value from AQ card
      RAW_MAX : Int := 27648;   // Raw maximum value from AQ card
   END_STRUCT;
END_TYPE

// folder: 10 - 19 IO & Processing

DATA_BLOCK "10 DI_DATA"   // DB10
TITLE = Digital Input Data
{ S7_Optimized_Access := 'TRUE' }
AUTHOR : JRS
VERSION : 0.1
// Processed data for code use
   VAR
      R2_SPR_DI_0_2 : Bool;   // Spare input
      R2_SPR_DI_0_3 : Bool;   // Spare input
      R2_SPR_DI_1_6 : Bool;   // Spare input
      R2_SPR_DI_3_2 : Bool;   // Spare input
      R2_SPR_DI_3_7 : Bool;   // Spare input
      ESD_OK : Bool;   // External shutdown
      S2_8K1_OK : Bool;   // IGG E-Stop healthy
      E131_WRNG : Bool;   // E131 I&A Air Compressor warning
      E131_OK : Bool;   // E131 I&A Air Compressor Running
      E131_SHTDN : Bool;   // E131 I&A Air Compressor Shut down
      E600_NOK : Bool;   // Oxygen Analyser E600 system fail
      E600_HIHI : Bool;   // Oxygen Analyser E600 high high setpoint
      E600_LOLO : Bool;   // Oxygen Analyser E600 low low
      E600_PWR_OK : Bool;   // Oxygen Analyser E600 power healthy
      E700_OPACITY : Bool;   // Soot Monitor E700 opacity
      E700_PWR_OK : Bool;   // Soot Monitor E700 Power Healthy
      FD001_OK : Bool;   // Flame Detector FD001 OK
      FD001_PWR_OK : Bool;   // Flame Detector FD001 Power Healthy
      FD001_FLAME_DETCTN : Bool;   // Flame Detector FD001 Flame Detect
      FS115 : Bool;   // Main atom air flow switch
      FS123 : Bool;   // Pilot ignition air flow switch
      FS317 : Bool;   // Jacket cooling water flow switch
      FS320 : Bool;   // Nozzle cooling water flow switch
      LS001 : Bool;   // Shell CW level hi hi switch
      P301_ENBLD : Bool;   // CSW Pump enabled
      P301_TRIPPED : Bool;   // CSW pump tripped
      P305_ENBLD : Bool;   // Fresh water pump enabled
      P305_TRIPPED : Bool;   // Fresh water pump tripped
      PS101 : Bool;   // CA pressure switch
      TS006 : Bool;   // IG Shell Temp Hi Switch
      TS403_FAULT : Bool;   // IG temp hi hi switch
      X001_PWR_OK : Bool;   // Ignitor Power Healthy
   END_VAR
BEGIN
END_DATA_BLOCK

DATA_BLOCK "12_AI_Data"   // DB12
TITLE = Analogue Input Data
{ S7_Optimized_Access := 'TRUE' }
AUTHOR : JRS
VERSION : 0.1
// Processed data for code use
   VAR
      PIT112In_SCALED : Real;   // IA Inlet pressure
      PIT205In_SCALED : Real;   // IGG Main fuel pressure
      FD001FlameSignalIn : Real;   // Flame signal
      PIT113In_SCALED : Real;   // IGG Main atom air pressure
      R2_SPR_AI_102_SCALED : Real;   // Spare input
      PIT204In_SCALED : Real;   // IGG Inlet fuel pressure
      TIT202In_SCALED : Real;   // IGG Inlet fuel temperature
      E600O2ContentIn : Real;   // O2 Analyser content
      E700SootContentIn : Real;   // IG Soot content
      IW_96 : "AI_Data";   // PIT205 calibration
      IW_98 : "AI_Data";   // FD001 calibration
      IW_100 : "AI_Data";   // PIT113 calibration data
      IW_102 : "AI_Data";   // PIT112 calibration data
      IW_104 : "AI_Data";   // PIT204 calibration data
      IW_106 : "AI_Data";   // TIT202 calibration data
      IW_108 : "AI_Data";   // E600 calibration data
      IW_110 : "AI_Data";   // E700 calibration data
   END_VAR
BEGIN
   IW_98.ENG_MAX := 100.0;
   IW_96.ENG_MAX := 40.0;   // Engineering units maximum value - bar(g)
   IW_100.ENG_MAX := 40.0;   // Engineering units maximum value -bar(g)
   IW_104.ENG_MAX := 40.0;   // Engineering units maximum value - bar(g)
   IW_106.ENG_MAX := 150.0;   // Engineering units maximum value - degC
   IW_102.ENG_MAX := 40.0;   // Engineering units maximum value - bar(g)
   IW_102.ENG_MIN := 0.0;   // Engineering units minimum value - bar(g)
   IW_106.ENG_MIN := 0.0;   // Engineering units minimum value - degC
   IW_108.ENG_MIN := 0.0;   // Engineering units minimum value - (% O2)
   IW_108.ENG_MAX := 25.0;   // Engineering units maximum value - (% O2)
   IW_110.ENG_MIN := 0.0;   // Engineering units minimum value - % Opacity
   IW_110.ENG_MAX := 100.0;   // Engineering units maximum value - % Opacity
   IW_110.RAW_MIN := 0;
   IW_110.RAW_MAX := 27648;
   // IW_96.ENG_MIN : Engineering units minimum value - bar(g)
   // IW_100.ENG_MIN : Engineering units minimum value - bar(g)
   // IW_104.ENG_MIN : Engineering units minimum value - bar(g)
END_DATA_BLOCK

DATA_BLOCK "14_DQ_Data"   // DB14
TITLE = Digital Output Data
{ S7_Optimized_Access := 'TRUE' }
AUTHOR : JRS
VERSION : 0.1
// Processed data for output via physical connection
   VAR
      "200CV127ControlOut" : Bool;   // Test pressure valve control
      "200CV124ControlOut" : Bool;   // Pilot B ignition air valve control
      "200CV215ControlOut" : Bool;   // Pilot B fuel valve 1 control
      "200CV216ControlOut" : Bool;   // Pilot B fuel valve 2 control
      "200CV114ControlOut" : Bool;   // Main B atom air valve control
      "200CV206ControlOut" : Bool;   // Main B fuel valve 1 control
      "200CV207ControlOut" : Bool;   // Main B fuel valve 2 control
      E131ControlOut : Bool := true;   // IA Compressor Control
      X001ControlOut : Bool;   // Igniter control
      P301ControlOut : Bool;   // CSW Pump control
      P305ControlOut : Bool;   // Fresh water pump control
      R2_SPR_DQ_1_3 : Bool;   // Spare output
      R2_SPR_DQ_1_4 : Bool;   // Spare output
      R2_SPR_DQ_1_5 : Bool;   // Spare output
      R2_SPR_DQ_1_6 : Bool;   // Spare output
      R2_SPR_DQ_1_2 : Bool;   // Spare output
      "IA Compressor RE" : TON_TIME;
      "IA Compressor RE_TP" : TP_TIME;
   END_VAR
BEGIN
END_DATA_BLOCK

DATA_BLOCK "16_AQ_Data"   // DB16
TITLE = Analogue Output Data
{ S7_Optimized_Access := 'TRUE' }
AUTHOR : JRS
VERSION : 0.1
// Processed data for output via physical connection
   VAR
      R2_SPR_AQ_96 : Real;   // Spare output
      R2_SPR_AQ_98 : Real;   // Spare output
   END_VAR
   VAR RETAIN
      CV203_CNTRL : Real;   // Main fuel reg Valve Control
      CV111_CNTRL : Real;   // Main Atom Air Reg Valve Control
   END_VAR
   VAR
      QW_96 : "AQ_Data";   // Spare output calibration data
      QW_98 : "AQ_Data";   // Spare output calibration data
      QW_100 : "AQ_Data";   // CV203 calibration data
      QW_102 : "AQ_Data";   // CV111 calibration data
   END_VAR
BEGIN
   QW_100.ENG_MIN := 0.0;   // Engineering units minimum value - %
   QW_100.ENG_MAX := 100.0;   // Engineering units maximum value - %
   QW_102.ENG_MIN := 0.0;   // Engineering units minimum value - %
   QW_102.ENG_MAX := 100.0;   // Engineering units maximum value - %
END_DATA_BLOCK

DATA_BLOCK "19_AUTO_CMNDS_Data"   // DB19
TITLE = Automatic Commands Data
{ S7_Optimized_Access := 'TRUE' }
AUTHOR : JRS
VERSION : 0.1
// Defined data for use prior to output processing
   VAR
      IG_FLM_Demand : Bool;   // 1 = Run, 0 = Not
      MAIN_FLM_Demand : Bool;   // 1 = Run, 0 = Not
      IG_PRG_Demand : Bool;   // 1 = Run, 0 = Not
      CV203_PID_MDLTG : Bool;   // 1 = Run, 0 = Not
      CV111_PID_MDLTG : Bool;   // 1 = Run, 0 = Not
      CV203_AQ_VAL : Real;   // Output value for ramp start
      CV203_RAMP_CNTRL : Bool;   // 1 = Run, 0 = Not
      INTO_CV203_RAMP_EDGE : Bool;   // Edge bit
      CV111_AQ_VAL : Real;   // Output value for initial state
   END_VAR
BEGIN
END_DATA_BLOCK

DATA_BLOCK "Evolving Setpoint_DB"   // DB107
{ S7_Optimized_Access := 'TRUE' }
VERSION : 0.1
// stored: InstanceOfName Evolving Setpoint
"Evolving Setpoint"
BEGIN
END_DATA_BLOCK

DATA_BLOCK "IDB_E131_Functioning Hours"   // DB131
{ S7_Optimized_Access := 'TRUE' }
VERSION : 0.1
// stored: InstanceOfName 64_Functioning Hours
"64_Functioning Hours"
BEGIN
END_DATA_BLOCK

// folder: 100 - 199 Automatic Sequencing

DATA_BLOCK "100_BC_AUTO_SEQ_DB"   // DB100
{ S7_Optimized_Access := 'TRUE' }
VERSION : 0.1
// stored: InstanceOfName 100_BC_AUTO_SEQ
"100_BC_AUTO_SEQ"
BEGIN
END_DATA_BLOCK

DATA_BLOCK "102_Pilot_Burner_DB"   // DB102
{ S7_Optimized_Access := 'TRUE' }
FAMILY : JRS
VERSION : 0.1
// stored: InstanceOfName 102_Pilot_Burner
"102_Pilot_Burner"
BEGIN
   IGNTR_DLY := T#1s;
   FV1_DLY := T#1s;
   FV2_3W_DLY := T#1s;
   FD_DLY := T#1s;
   IGNTR_MAX_RT := T#20s;
END_DATA_BLOCK

DATA_BLOCK "103_Main_Burner_DB"   // DB103
{ S7_Optimized_Access := 'TRUE' }
AUTHOR : JRS
VERSION : 0.1
// stored: InstanceOfName 103_Main_Burner
"103_Main_Burner"
BEGIN
END_DATA_BLOCK

DATA_BLOCK "104_Pilot_Purge_DB"   // DB104
{ S7_Optimized_Access := 'TRUE' }
AUTHOR : JRS
VERSION : 0.1
// stored: InstanceOfName 104_Pilot_Purge
"104_Pilot_Purge"
BEGIN
END_DATA_BLOCK

DATA_BLOCK "106_O2_RAMP_CNTRL_DB"   // DB106
{ S7_Optimized_Access := 'TRUE' }
AUTHOR : JRS
VERSION : 0.1
// stored: InstanceOfName 106_O2_RAMP_CNTRL
"106_O2_RAMP_CNTRL"
BEGIN
END_DATA_BLOCK

// folder: 300 - 499 Counter and Timer DBs

DATA_BLOCK "300_AUT_SEQ_TMRS_DB"   // DB300
TITLE = Auto Sequence Timers Data
{ S7_Optimized_Access := 'TRUE' }
AUTHOR : JRS
VERSION : 0.1
// Data area for auto sequence timers
   VAR
      "CV127 Open Delay #1" : TON_TIME;   // Valve open for time #1
      "CV127 Closed Delay #1" : TON_TIME;   // Valve closed time
      "CV127 Open Delay #2" : TON_TIME;   // Valve open for time #2
      "CV127 Closed Delay #2" : TON_TIME;   // Valve closed time
      "CV124 Open Delay" : TON_TIME;   // Valve max move time, no tell back
      "CV114 Open Delay" : TON_TIME;   // Valve max move time, no tell back
      "CV206 Close Delay" : TON_TIME;   // Valve max move time, no tell back
      "CV207 Close Delay" : TON_TIME;   // Valve max move time, no tell back
      "CV114 Close Delay" : TON_TIME;   // Valve max move time, no tell back
      "CV215 Close Delay" : TON_TIME;   // Valve max move time, no tell back
      "CV216 Close Delay" : TON_TIME;   // Valve max move time, no tell back
      "CV124 Close Delay" : TON_TIME;   // Valve max move time, no tell back
      "CV127 Delay after Open" : TON_TIME;
      "FS317 Unhealthy Delay" : TON_TIME;
      "FS320 Unhealthy Delay" : TON_TIME;
      "CV111 After Open Delay" : TON_TIME;
      "PS111 Alarm Delay" : TON_TIME;
      "ALARM STOP TP" : TP_TIME;
      "Shutting down confirmed" : TP_TIME;
      "Modulation Stopped Confirmation To IGG" : TP_TIME;
      PILOT_PURGE_DN : TOF_TIME;
      "Pilot Flame Purge Sequence Failure" : TP_TIME;
      "P301 Delay after Start" : TON_TIME;
      SFTY_SYS_IL : TOF_TIME;
      "CV401 Not Closed Brake" : TON_TIME;
   END_VAR
BEGIN
   "CV127 Open Delay #1".PT := T#10s;
   "CV127 Delay after Open".PT := T#3s;
   "ALARM STOP TP".PT := T#1s;
   SFTY_SYS_IL.PT := T#1s;
   "CV401 Not Closed Brake".PT := T#10s;
END_DATA_BLOCK

// folder: 50 - 59 PLC Communication

DATA_BLOCK "50_CMND_DATA"   // DB50
TITLE = Command Data
{ S7_Optimized_Access := 'FALSE' }
AUTHOR : JRS